// TIA Portal project "Projekt_Serhii_Bodnia" (V19) (continued)

   FOR #forVal := 0 TO 120 DO
       FOR #forVal_2:=0 TO 10 DO
           #rdTimeReturn:=RD_SYS_T(#outputTime);
           #rdTimeReturn := WR_SYS_T(#outputTime);
           #rdTimeReturn := RD_SYS_T(#outputTime);
           #rdTimeReturn := WR_SYS_T(#outputTime);
       END_FOR;
       #SyncVal:= PEEK(area := 16#81,
                      dbNumber := 0,
                      byteOffset := 511);
       IF #SyncVal = #CompVal THEN
          GOTO M_1;
       END_IF;
   END_FOR;
   RETURN;

   M_1:
   POKE(area := 16#81,
        dbNumber := 0,
        byteOffset := 511,
        value := B#16#0);
END_FUNCTION

ORGANIZATION_BLOCK "Main"   // OB1, FBD, ProgramCycle
TITLE = "Main Program Sweep (Cycle)"
{ S7_Optimized_Access := 'TRUE' }
VERSION : 0.1
   VAR_INPUT
      Initial_Call : Bool;   // Initial call of this OB
      Remanence : Bool;   // =True, if remanent data are available
   END_VAR
BEGIN

REGION Network 1: Konnektierungsbaustein für PLC-Lab / Factory IO
   // Im Netzwerk 1 wird der Konnektierungsbaustein für PLC-Lab aufgerufen.
   // Dieser Aufruf darf nicht entfernt werden!
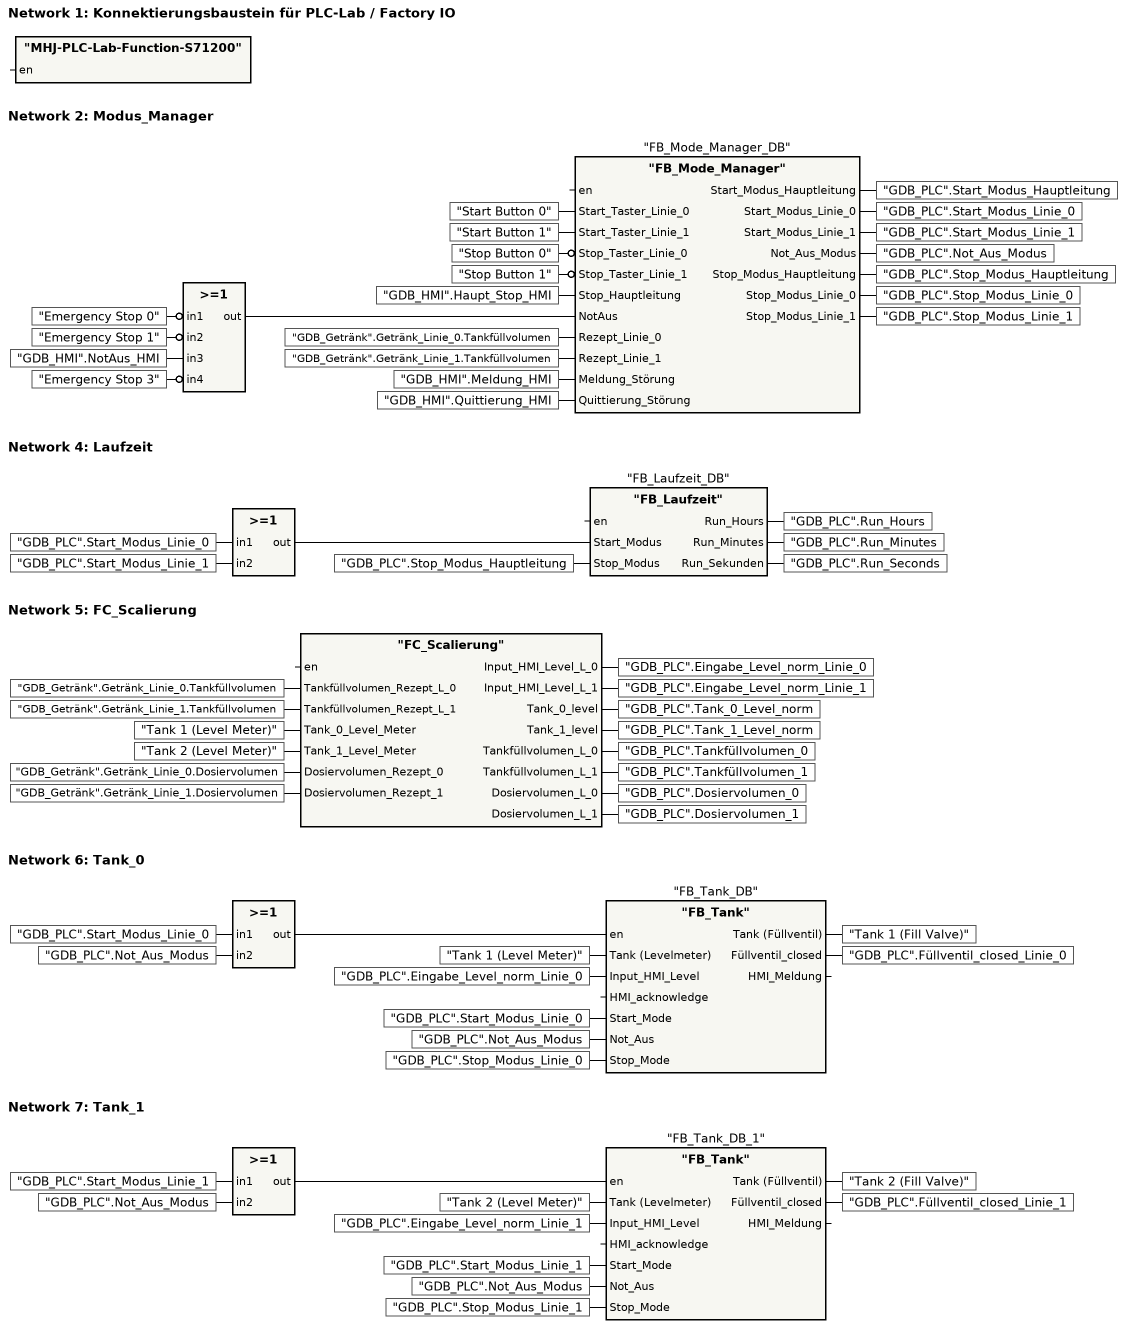
   "MHJ-PLC-Lab-Function-S71200"();
END_REGION

REGION Network 2: Modus_Manager
   "FB_Mode_Manager_DB"(Start_Taster_Linie_0 := "Start Button 0",   // "FB_Mode_Manager"
                        Start_Taster_Linie_1 := "Start Button 1",
                        Stop_Taster_Linie_0 := NOT "Stop Button 0",
                        Stop_Taster_Linie_1 := NOT "Stop Button 1",
                        Stop_Hauptleitung := "GDB_HMI".Haupt_Stop_HMI,
                        NotAus := NOT "Emergency Stop 0" OR NOT "Emergency Stop 1" OR "GDB_HMI".NotAus_HMI OR NOT "Emergency Stop 3",
                        Rezept_Linie_0 := "GDB_Getränk".Getränk_Linie_0.Tankfüllvolumen,
                        Rezept_Linie_1 := "GDB_Getränk".Getränk_Linie_1.Tankfüllvolumen,
                        Meldung_Störung := "GDB_HMI".Meldung_HMI,
                        Quittierung_Störung := "GDB_HMI".Quittierung_HMI,
                        Start_Modus_Hauptleitung => "GDB_PLC".Start_Modus_Hauptleitung,
                        Start_Modus_Linie_0 => "GDB_PLC".Start_Modus_Linie_0,
                        Start_Modus_Linie_1 => "GDB_PLC".Start_Modus_Linie_1,
                        Not_Aus_Modus => "GDB_PLC".Not_Aus_Modus,
                        Stop_Modus_Hauptleitung => "GDB_PLC".Stop_Modus_Hauptleitung,
                        Stop_Modus_Linie_0 => "GDB_PLC".Stop_Modus_Linie_0,
                        Stop_Modus_Linie_1 => "GDB_PLC".Stop_Modus_Linie_1);
END_REGION

REGION Network 3 (SCL): Störung Meldungen
   "GDB_PLC".Störung[0] := "GDB_HMI".Meldung_HMI.%X0;
   "GDB_PLC".Störung[1] := "GDB_HMI".Meldung_HMI.%X1;
   "GDB_PLC".Störung[2] := "GDB_HMI".Meldung_HMI.%X2;
   "GDB_PLC".Störung[3] := "GDB_HMI".Meldung_HMI.%X3;
   "GDB_PLC".Störung[4] := "GDB_HMI".Meldung_HMI.%X4;
   "GDB_PLC".Störung[5] := "GDB_HMI".Meldung_HMI.%X5;
   "GDB_PLC".Störung[6] := "GDB_HMI".Meldung_HMI.%X6;
   "GDB_PLC".Störung[7] := "GDB_HMI".Meldung_HMI.%X7;
   "GDB_PLC".Störung[8] := "GDB_HMI".Meldung_HMI.%X8;
   "GDB_PLC".Störung[9] := "GDB_HMI".Meldung_HMI.%X9;
   "GDB_PLC".Störung[10] := "GDB_HMI".Meldung_HMI.%X10;
   "GDB_PLC".Störung[11] := "GDB_HMI".Meldung_HMI.%X11;
   "GDB_PLC".Störung[12] := "GDB_HMI".Meldung_HMI.%X12;
   "GDB_PLC".Störung[13] := "GDB_HMI".Meldung_HMI.%X13;
   "GDB_PLC".Störung[14] := "GDB_HMI".Meldung_HMI.%X14;
   "GDB_PLC".Störung[15] := "GDB_HMI".Meldung_HMI.%X15;
END_REGION

REGION Network 4: Laufzeit
   "FB_Laufzeit_DB"(Start_Modus := "GDB_PLC".Start_Modus_Linie_0 OR "GDB_PLC".Start_Modus_Linie_1,   // "FB_Laufzeit"
                    Stop_Modus := "GDB_PLC".Stop_Modus_Hauptleitung,
                    Run_Hours => "GDB_PLC".Run_Hours,
                    Run_Minutes => "GDB_PLC".Run_Minutes,
                    Run_Sekunden => "GDB_PLC".Run_Seconds);
END_REGION

REGION Network 5: FC_Scalierung
   "FC_Scalierung"(Tankfüllvolumen_Rezept_L_0 := "GDB_Getränk".Getränk_Linie_0.Tankfüllvolumen,
                   Tankfüllvolumen_Rezept_L_1 := "GDB_Getränk".Getränk_Linie_1.Tankfüllvolumen,
                   Tank_0_Level_Meter := "Tank 1 (Level Meter)",
                   Tank_1_Level_Meter := "Tank 2 (Level Meter)",
                   Dosiervolumen_Rezept_0 := "GDB_Getränk".Getränk_Linie_0.Dosiervolumen,
                   Dosiervolumen_Rezept_1 := "GDB_Getränk".Getränk_Linie_1.Dosiervolumen,
                   Input_HMI_Level_L_0 => "GDB_PLC".Eingabe_Level_norm_Linie_0,
                   Input_HMI_Level_L_1 => "GDB_PLC".Eingabe_Level_norm_Linie_1,
                   Tank_0_level => "GDB_PLC".Tank_0_Level_norm,
                   Tank_1_level => "GDB_PLC".Tank_1_Level_norm,
                   Tankfüllvolumen_L_0 => "GDB_PLC".Tankfüllvolumen_0,
                   Tankfüllvolumen_L_1 => "GDB_PLC".Tankfüllvolumen_1,
                   Dosiervolumen_L_0 => "GDB_PLC".Dosiervolumen_0,
                   Dosiervolumen_L_1 => "GDB_PLC".Dosiervolumen_1);
END_REGION

REGION Network 6: Tank_0
   IF "GDB_PLC".Start_Modus_Linie_0 OR "GDB_PLC".Not_Aus_Modus THEN
       "FB_Tank_DB"("Tank (Levelmeter)" := "Tank 1 (Level Meter)",   // "FB_Tank"
                    Input_HMI_Level := "GDB_PLC".Eingabe_Level_norm_Linie_0,
                    Start_Mode := "GDB_PLC".Start_Modus_Linie_0,
                    Not_Aus := "GDB_PLC".Not_Aus_Modus,
                    Stop_Mode := "GDB_PLC".Stop_Modus_Linie_0,
                    "Tank (Füllventil)" => "Tank 1 (Fill Valve)",
                    Füllventil_closed => "GDB_PLC".Füllventil_closed_Linie_0);
   END_IF;
END_REGION

REGION Network 7: Tank_1
   IF "GDB_PLC".Start_Modus_Linie_1 OR "GDB_PLC".Not_Aus_Modus THEN
       "FB_Tank_DB_1"("Tank (Levelmeter)" := "Tank 2 (Level Meter)",   // "FB_Tank"
                      Input_HMI_Level := "GDB_PLC".Eingabe_Level_norm_Linie_1,
                      Start_Mode := "GDB_PLC".Start_Modus_Linie_1,
                      Not_Aus := "GDB_PLC".Not_Aus_Modus,
                      Stop_Mode := "GDB_PLC".Stop_Modus_Linie_1,
                      "Tank (Füllventil)" => "Tank 2 (Fill Valve)",
                      Füllventil_closed => "GDB_PLC".Füllventil_closed_Linie_1);
   END_IF;
END_REGION

REGION Network 8: Abfüllmaschine_Band_0
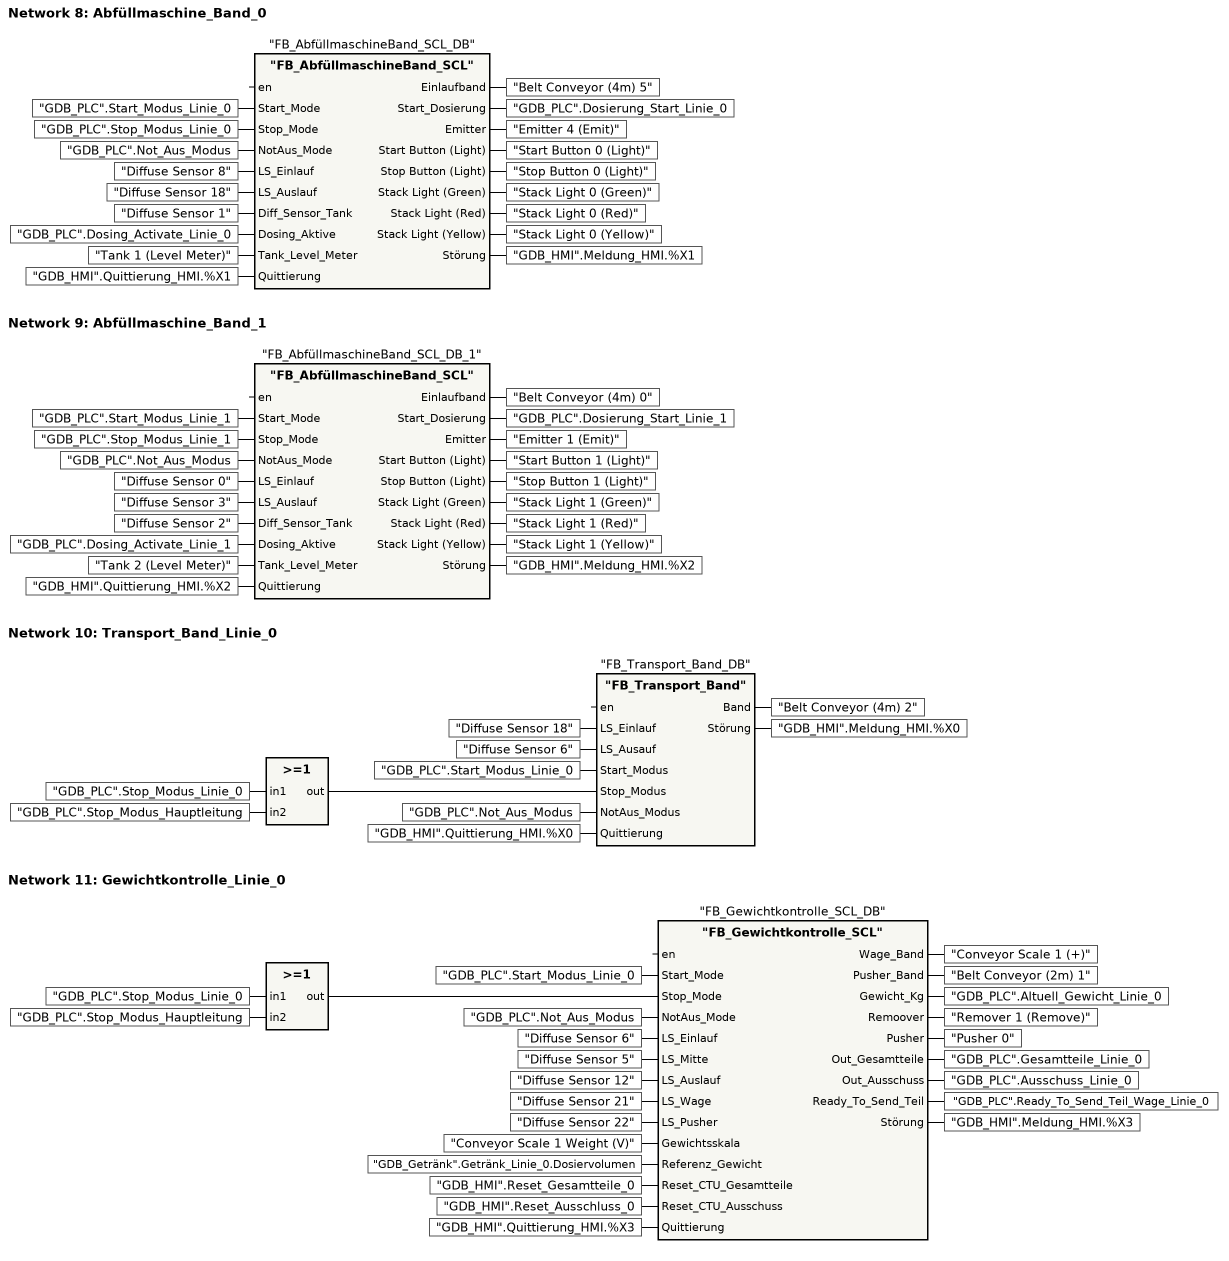
   "FB_AbfüllmaschineBand_SCL_DB"(Start_Mode := "GDB_PLC".Start_Modus_Linie_0,   // "FB_AbfüllmaschineBand_SCL"
                           Stop_Mode := "GDB_PLC".Stop_Modus_Linie_0,
                           NotAus_Mode := "GDB_PLC".Not_Aus_Modus,
                           LS_Einlauf := "Diffuse Sensor 8",
                           LS_Auslauf := "Diffuse Sensor 18",
                           Diff_Sensor_Tank := "Diffuse Sensor 1",
                           Dosing_Aktive := "GDB_PLC".Dosing_Activate_Linie_0,
                           Tank_Level_Meter := "Tank 1 (Level Meter)",
                           Quittierung := "GDB_HMI".Quittierung_HMI.%X1,
                           Einlaufband => "Belt Conveyor (4m) 5",
                           Start_Dosierung => "GDB_PLC".Dosierung_Start_Linie_0,
                           Emitter => "Emitter 4 (Emit)",
                           "Start Button (Light)" => "Start Button 0 (Light)",
                           "Stop Button (Light)" => "Stop Button 0 (Light)",
                           "Stack Light (Green)" => "Stack Light 0 (Green)",
                           "Stack Light (Red)" => "Stack Light 0 (Red)",
                           "Stack Light (Yellow)" => "Stack Light 0 (Yellow)",
                           Störung => "GDB_HMI".Meldung_HMI.%X1);
END_REGION

REGION Network 9: Abfüllmaschine_Band_1
   "FB_AbfüllmaschineBand_SCL_DB_1"(Start_Mode := "GDB_PLC".Start_Modus_Linie_1,   // "FB_AbfüllmaschineBand_SCL"
                           Stop_Mode := "GDB_PLC".Stop_Modus_Linie_1,
                           NotAus_Mode := "GDB_PLC".Not_Aus_Modus,
                           LS_Einlauf := "Diffuse Sensor 0",
                           LS_Auslauf := "Diffuse Sensor 3",
                           Diff_Sensor_Tank := "Diffuse Sensor 2",
                           Dosing_Aktive := "GDB_PLC".Dosing_Activate_Linie_1,
                           Tank_Level_Meter := "Tank 2 (Level Meter)",
                           Quittierung := "GDB_HMI".Quittierung_HMI.%X2,
                           Einlaufband => "Belt Conveyor (4m) 0",
                           Start_Dosierung => "GDB_PLC".Dosierung_Start_Linie_1,
                           Emitter => "Emitter 1 (Emit)",
                           "Start Button (Light)" => "Start Button 1 (Light)",
                           "Stop Button (Light)" => "Stop Button 1 (Light)",
                           "Stack Light (Green)" => "Stack Light 1 (Green)",
                           "Stack Light (Red)" => "Stack Light 1 (Red)",
                           "Stack Light (Yellow)" => "Stack Light 1 (Yellow)",
                           Störung => "GDB_HMI".Meldung_HMI.%X2);
END_REGION

REGION Network 10: Transport_Band_Linie_0
   "FB_Transport_Band_DB"(LS_Einlauf := "Diffuse Sensor 18",   // "FB_Transport_Band"
                          LS_Ausauf := "Diffuse Sensor 6",
                          Start_Modus := "GDB_PLC".Start_Modus_Linie_0,
                          Stop_Modus := "GDB_PLC".Stop_Modus_Linie_0 OR "GDB_PLC".Stop_Modus_Hauptleitung,
                          NotAus_Modus := "GDB_PLC".Not_Aus_Modus,
                          Quittierung := "GDB_HMI".Quittierung_HMI.%X0,
                          Band => "Belt Conveyor (4m) 2",
                          Störung => "GDB_HMI".Meldung_HMI.%X0);
END_REGION

REGION Network 11: Gewichtkontrolle_Linie_0
   "FB_Gewichtkontrolle_SCL_DB"(Start_Mode := "GDB_PLC".Start_Modus_Linie_0,   // "FB_Gewichtkontrolle_SCL"
                           Stop_Mode := "GDB_PLC".Stop_Modus_Linie_0 OR "GDB_PLC".Stop_Modus_Hauptleitung,
                           NotAus_Mode := "GDB_PLC".Not_Aus_Modus,
                           LS_Einlauf := "Diffuse Sensor 6",
                           LS_Mitte := "Diffuse Sensor 5",
                           LS_Auslauf := "Diffuse Sensor 12",
                           LS_Wage := "Diffuse Sensor 21",
                           LS_Pusher := "Diffuse Sensor 22",
                           Gewichtsskala := "Conveyor Scale 1 Weight (V)",
                           Referenz_Gewicht := "GDB_Getränk".Getränk_Linie_0.Dosiervolumen,
                           Reset_CTU_Gesamtteile := "GDB_HMI".Reset_Gesamtteile_0,
                           Reset_CTU_Ausschuss := "GDB_HMI".Reset_Ausschluss_0,
                           Quittierung := "GDB_HMI".Quittierung_HMI.%X3,
                           Wage_Band => "Conveyor Scale 1 (+)",
                           Pusher_Band => "Belt Conveyor (2m) 1",
                           Gewicht_Kg => "GDB_PLC".Altuell_Gewicht_Linie_0,
                           Remoover => "Remover 1 (Remove)",
                           Pusher => "Pusher 0",
                           Out_Gesamtteile => "GDB_PLC".Gesamtteile_Linie_0,
                           Out_Ausschuss => "GDB_PLC".Ausschuss_Linie_0,
                           Ready_To_Send_Teil => "GDB_PLC".Ready_To_Send_Teil_Wage_Linie_0,
                           Störung => "GDB_HMI".Meldung_HMI.%X3);
END_REGION

REGION Network 12: Gewichtkontrolle_Linie_1
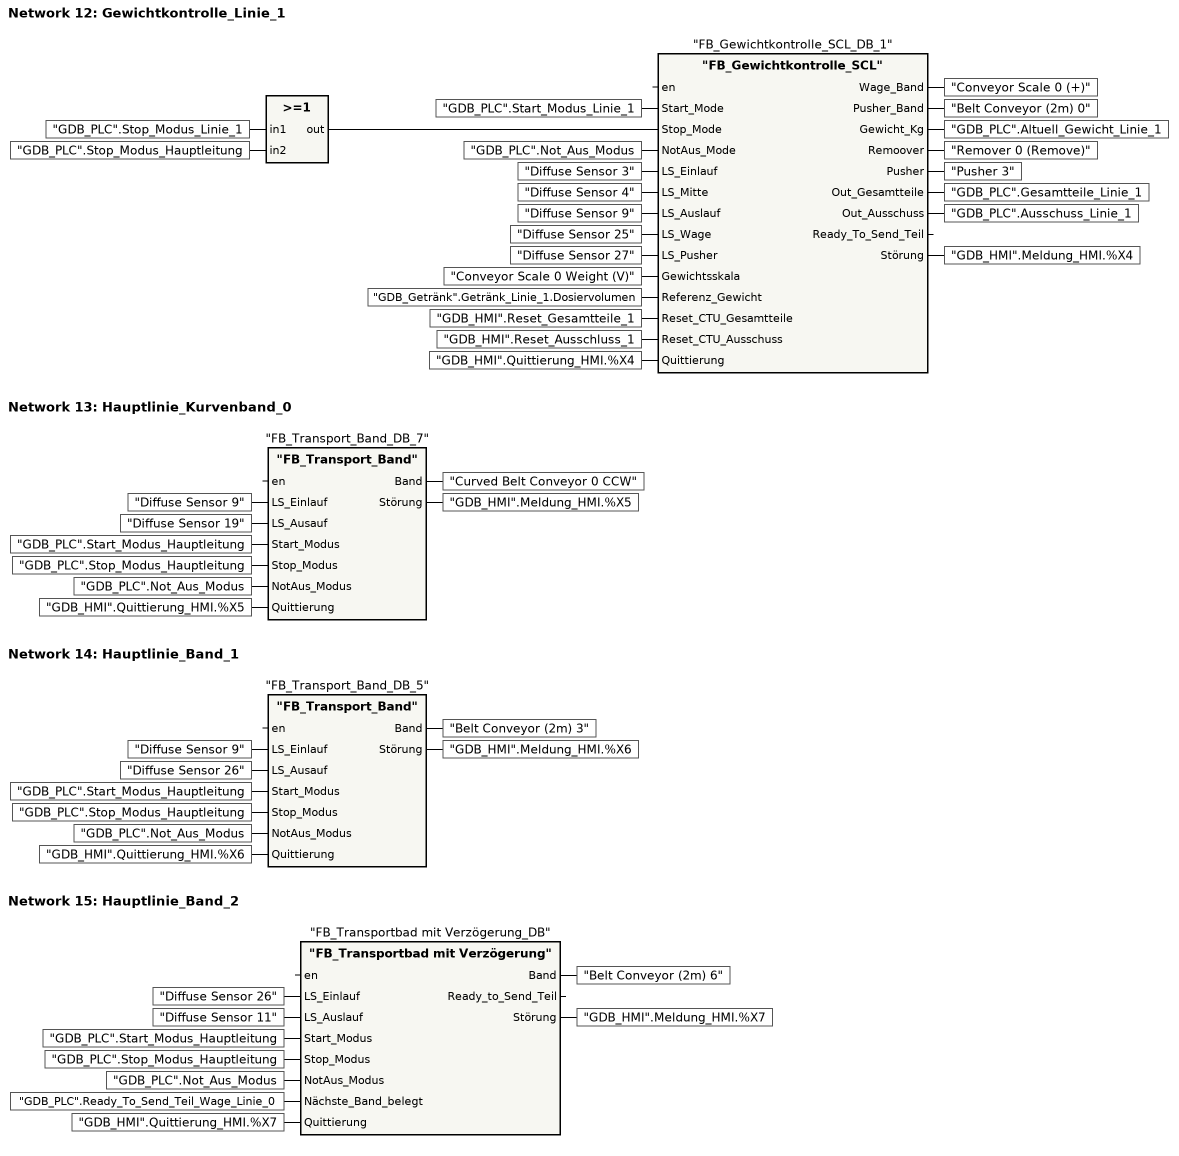
   "FB_Gewichtkontrolle_SCL_DB_1"(Start_Mode := "GDB_PLC".Start_Modus_Linie_1,   // "FB_Gewichtkontrolle_SCL"
                           Stop_Mode := "GDB_PLC".Stop_Modus_Linie_1 OR "GDB_PLC".Stop_Modus_Hauptleitung,
                           NotAus_Mode := "GDB_PLC".Not_Aus_Modus,
                           LS_Einlauf := "Diffuse Sensor 3",
                           LS_Mitte := "Diffuse Sensor 4",
                           LS_Auslauf := "Diffuse Sensor 9",
                           LS_Wage := "Diffuse Sensor 25",
                           LS_Pusher := "Diffuse Sensor 27",
                           Gewichtsskala := "Conveyor Scale 0 Weight (V)",
                           Referenz_Gewicht := "GDB_Getränk".Getränk_Linie_1.Dosiervolumen,
                           Reset_CTU_Gesamtteile := "GDB_HMI".Reset_Gesamtteile_1,
                           Reset_CTU_Ausschuss := "GDB_HMI".Reset_Ausschluss_1,
                           Quittierung := "GDB_HMI".Quittierung_HMI.%X4,
                           Wage_Band => "Conveyor Scale 0 (+)",
                           Pusher_Band => "Belt Conveyor (2m) 0",
                           Gewicht_Kg => "GDB_PLC".Altuell_Gewicht_Linie_1,
                           Remoover => "Remover 0 (Remove)",
                           Pusher => "Pusher 3",
                           Out_Gesamtteile => "GDB_PLC".Gesamtteile_Linie_1,
                           Out_Ausschuss => "GDB_PLC".Ausschuss_Linie_1,
                           Störung => "GDB_HMI".Meldung_HMI.%X4);
END_REGION

REGION Network 13: Hauptlinie_Kurvenband_0
   "FB_Transport_Band_DB_7"(LS_Einlauf := "Diffuse Sensor 9",   // "FB_Transport_Band"
                           LS_Ausauf := "Diffuse Sensor 19",
                           Start_Modus := "GDB_PLC".Start_Modus_Hauptleitung,
                           Stop_Modus := "GDB_PLC".Stop_Modus_Hauptleitung,
                           NotAus_Modus := "GDB_PLC".Not_Aus_Modus,
                           Quittierung := "GDB_HMI".Quittierung_HMI.%X5,
                           Band => "Curved Belt Conveyor 0 CCW",
                           Störung => "GDB_HMI".Meldung_HMI.%X5);
END_REGION

REGION Network 14: Hauptlinie_Band_1
   "FB_Transport_Band_DB_5"(LS_Einlauf := "Diffuse Sensor 9",   // "FB_Transport_Band"
                           LS_Ausauf := "Diffuse Sensor 26",
                           Start_Modus := "GDB_PLC".Start_Modus_Hauptleitung,
                           Stop_Modus := "GDB_PLC".Stop_Modus_Hauptleitung,
                           NotAus_Modus := "GDB_PLC".Not_Aus_Modus,
                           Quittierung := "GDB_HMI".Quittierung_HMI.%X6,
                           Band => "Belt Conveyor (2m) 3",
                           Störung => "GDB_HMI".Meldung_HMI.%X6);
END_REGION

REGION Network 15: Hauptlinie_Band_2
   "FB_Transportbad mit Verzögerung_DB"(LS_Einlauf := "Diffuse Sensor 26",   // "FB_Transportbad mit Verzögerung"
                           LS_Auslauf := "Diffuse Sensor 11",
                           Start_Modus := "GDB_PLC".Start_Modus_Hauptleitung,
                           Stop_Modus := "GDB_PLC".Stop_Modus_Hauptleitung,
                           NotAus_Modus := "GDB_PLC".Not_Aus_Modus,
                           Nächste_Band_belegt := "GDB_PLC".Ready_To_Send_Teil_Wage_Linie_0,
                           Quittierung := "GDB_HMI".Quittierung_HMI.%X7,
                           Band => "Belt Conveyor (2m) 6",
                           Störung => "GDB_HMI".Meldung_HMI.%X7);
END_REGION

REGION Network 16: Hauptlinie_T - Band_3
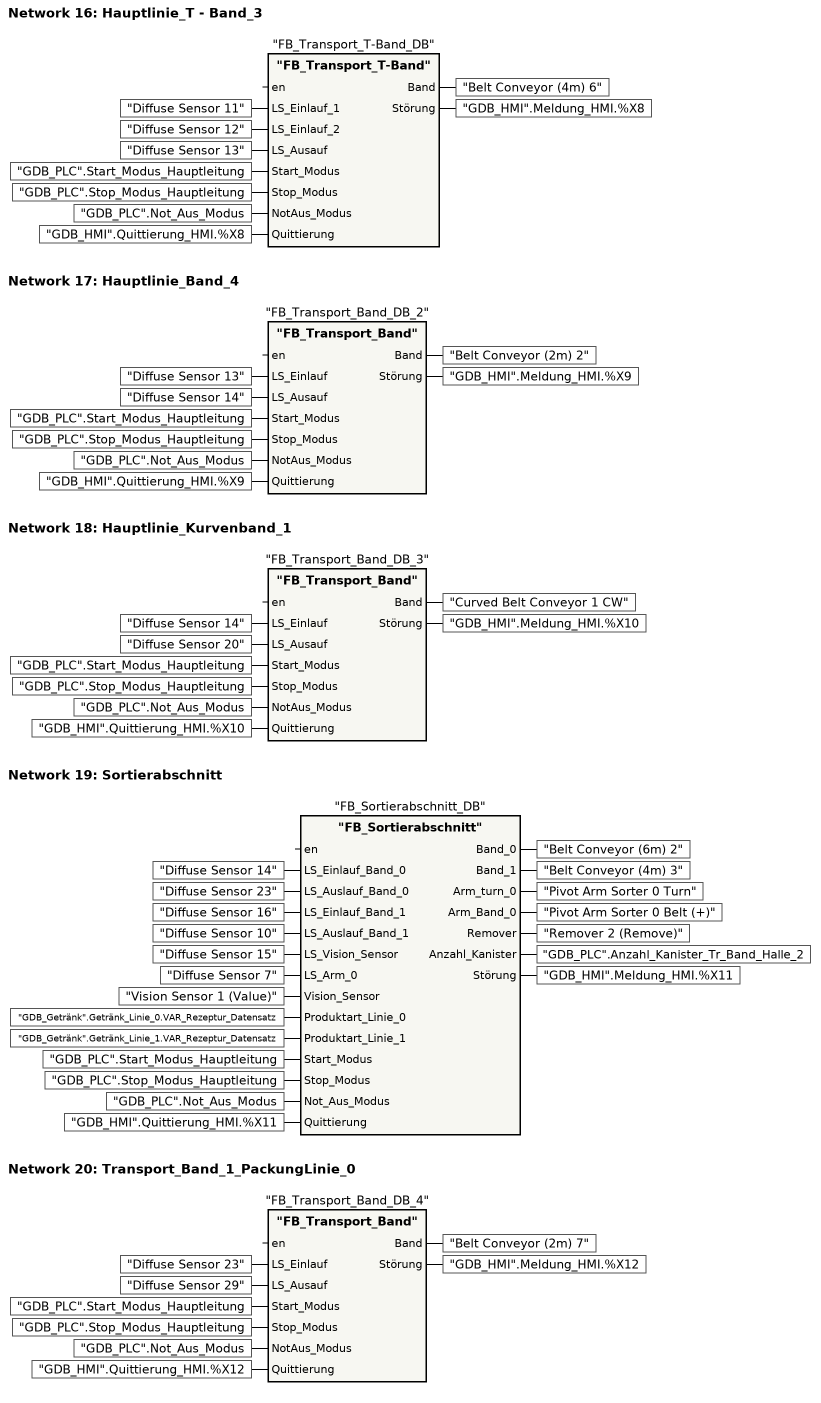
   "FB_Transport_T-Band_DB"(LS_Einlauf_1 := "Diffuse Sensor 11",   // "FB_Transport_T-Band"
                           LS_Einlauf_2 := "Diffuse Sensor 12",
                           LS_Ausauf := "Diffuse Sensor 13",
                           Start_Modus := "GDB_PLC".Start_Modus_Hauptleitung,
                           Stop_Modus := "GDB_PLC".Stop_Modus_Hauptleitung,
                           NotAus_Modus := "GDB_PLC".Not_Aus_Modus,
                           Quittierung := "GDB_HMI".Quittierung_HMI.%X8,
                           Band => "Belt Conveyor (4m) 6",
                           Störung => "GDB_HMI".Meldung_HMI.%X8);
END_REGION

REGION Network 17: Hauptlinie_Band_4
   "FB_Transport_Band_DB_2"(LS_Einlauf := "Diffuse Sensor 13",   // "FB_Transport_Band"
                           LS_Ausauf := "Diffuse Sensor 14",
                           Start_Modus := "GDB_PLC".Start_Modus_Hauptleitung,
                           Stop_Modus := "GDB_PLC".Stop_Modus_Hauptleitung,
                           NotAus_Modus := "GDB_PLC".Not_Aus_Modus,
                           Quittierung := "GDB_HMI".Quittierung_HMI.%X9,
                           Band => "Belt Conveyor (2m) 2",
                           Störung => "GDB_HMI".Meldung_HMI.%X9);
END_REGION

REGION Network 18: Hauptlinie_Kurvenband_1
   "FB_Transport_Band_DB_3"(LS_Einlauf := "Diffuse Sensor 14",   // "FB_Transport_Band"
                           LS_Ausauf := "Diffuse Sensor 20",
                           Start_Modus := "GDB_PLC".Start_Modus_Hauptleitung,
                           Stop_Modus := "GDB_PLC".Stop_Modus_Hauptleitung,
                           NotAus_Modus := "GDB_PLC".Not_Aus_Modus,
                           Quittierung := "GDB_HMI".Quittierung_HMI.%X10,
                           Band => "Curved Belt Conveyor 1 CW",
                           Störung => "GDB_HMI".Meldung_HMI.%X10);
END_REGION

REGION Network 19: Sortierabschnitt
   "FB_Sortierabschnitt_DB"(LS_Einlauf_Band_0 := "Diffuse Sensor 14",   // "FB_Sortierabschnitt"
                           LS_Auslauf_Band_0 := "Diffuse Sensor 23",
                           LS_Einlauf_Band_1 := "Diffuse Sensor 16",
                           LS_Auslauf_Band_1 := "Diffuse Sensor 10",
                           LS_Vision_Sensor := "Diffuse Sensor 15",
                           LS_Arm_0 := "Diffuse Sensor 7",
                           Vision_Sensor := "Vision Sensor 1 (Value)",
                           Produktart_Linie_0 := "GDB_Getränk".Getränk_Linie_0.VAR_Rezeptur_Datensatz,
                           Produktart_Linie_1 := "GDB_Getränk".Getränk_Linie_1.VAR_Rezeptur_Datensatz,
                           Start_Modus := "GDB_PLC".Start_Modus_Hauptleitung,
                           Stop_Modus := "GDB_PLC".Stop_Modus_Hauptleitung,
                           Not_Aus_Modus := "GDB_PLC".Not_Aus_Modus,
                           Quittierung := "GDB_HMI".Quittierung_HMI.%X11,
                           Band_0 => "Belt Conveyor (6m) 2",
                           Band_1 => "Belt Conveyor (4m) 3",
                           Arm_turn_0 => "Pivot Arm Sorter 0 Turn",
                           Arm_Band_0 => "Pivot Arm Sorter 0 Belt (+)",
                           Remover => "Remover 2 (Remove)",
                           Anzahl_Kanister => "GDB_PLC".Anzahl_Kanister_Tr_Band_Halle_2,
                           Störung => "GDB_HMI".Meldung_HMI.%X11);
END_REGION

REGION Network 20: Transport_Band_1_PackungLinie_0
   "FB_Transport_Band_DB_4"(LS_Einlauf := "Diffuse Sensor 23",   // "FB_Transport_Band"
                           LS_Ausauf := "Diffuse Sensor 29",
                           Start_Modus := "GDB_PLC".Start_Modus_Hauptleitung,
                           Stop_Modus := "GDB_PLC".Stop_Modus_Hauptleitung,
                           NotAus_Modus := "GDB_PLC".Not_Aus_Modus,
                           Quittierung := "GDB_HMI".Quittierung_HMI.%X12,
                           Band => "Belt Conveyor (2m) 7",
                           Störung => "GDB_HMI".Meldung_HMI.%X12);
END_REGION

REGION Network 21: Transport_Band_2_PackungLinie_0
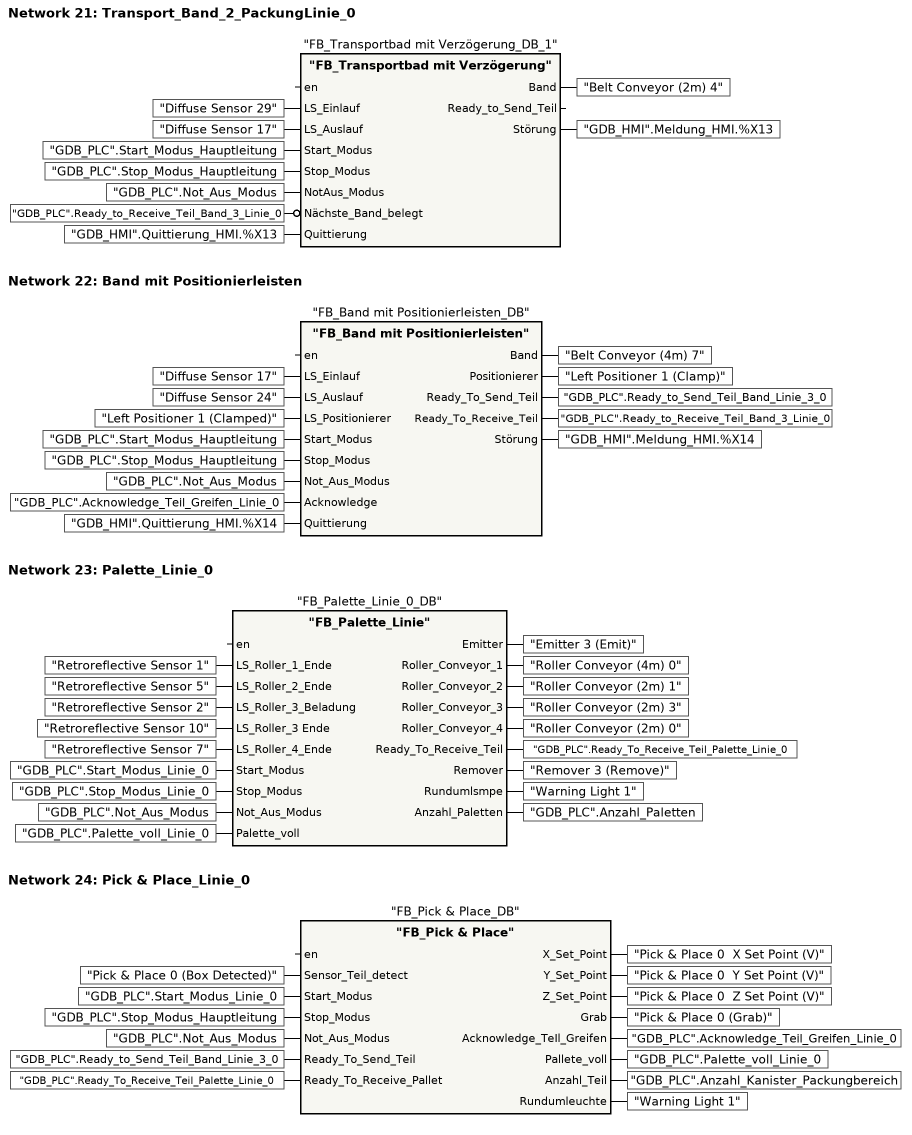
   "FB_Transportbad mit Verzögerung_DB_1"(LS_Einlauf := "Diffuse Sensor 29",   // "FB_Transportbad mit Verzögerung"
                           LS_Auslauf := "Diffuse Sensor 17",
                           Start_Modus := "GDB_PLC".Start_Modus_Hauptleitung,
                           Stop_Modus := "GDB_PLC".Stop_Modus_Hauptleitung,
                           NotAus_Modus := "GDB_PLC".Not_Aus_Modus,
                           Nächste_Band_belegt := NOT "GDB_PLC".Ready_to_Receive_Teil_Band_3_Linie_0,
                           Quittierung := "GDB_HMI".Quittierung_HMI.%X13,
                           Band => "Belt Conveyor (2m) 4",
                           Störung => "GDB_HMI".Meldung_HMI.%X13);
END_REGION

REGION Network 22: Band mit Positionierleisten
   "FB_Band mit Positionierleisten_DB"(LS_Einlauf := "Diffuse Sensor 17",   // "FB_Band mit Positionierleisten"
                           LS_Auslauf := "Diffuse Sensor 24",
                           LS_Positionierer := "Left Positioner 1 (Clamped)",
                           Start_Modus := "GDB_PLC".Start_Modus_Hauptleitung,
                           Stop_Modus := "GDB_PLC".Stop_Modus_Hauptleitung,
                           Not_Aus_Modus := "GDB_PLC".Not_Aus_Modus,
                           Acknowledge := "GDB_PLC".Acknowledge_Teil_Greifen_Linie_0,
                           Quittierung := "GDB_HMI".Quittierung_HMI.%X14,
                           Band => "Belt Conveyor (4m) 7",
                           Positionierer => "Left Positioner 1 (Clamp)",
                           Ready_To_Send_Teil => "GDB_PLC".Ready_to_Send_Teil_Band_Linie_3_0,
                           Ready_To_Receive_Teil => "GDB_PLC".Ready_to_Receive_Teil_Band_3_Linie_0,
                           Störung => "GDB_HMI".Meldung_HMI.%X14);
END_REGION

REGION Network 23: Palette_Linie_0
   "FB_Palette_Linie_0_DB"(LS_Roller_1_Ende := "Retroreflective Sensor 1",   // "FB_Palette_Linie"
                           LS_Roller_2_Ende := "Retroreflective Sensor 5",
                           LS_Roller_3_Beladung := "Retroreflective Sensor 2",
                           "LS_Roller_3 Ende" := "Retroreflective Sensor 10",
                           LS_Roller_4_Ende := "Retroreflective Sensor 7",
                           Start_Modus := "GDB_PLC".Start_Modus_Linie_0,
                           Stop_Modus := "GDB_PLC".Stop_Modus_Linie_0,
                           Not_Aus_Modus := "GDB_PLC".Not_Aus_Modus,
                           Palette_voll := "GDB_PLC".Palette_voll_Linie_0,
                           Emitter => "Emitter 3 (Emit)",
                           Roller_Conveyor_1 => "Roller Conveyor (4m) 0",
                           Roller_Conveyor_2 => "Roller Conveyor (2m) 1",
                           Roller_Conveyor_3 => "Roller Conveyor (2m) 3",
                           Roller_Conveyor_4 => "Roller Conveyor (2m) 0",
                           Ready_To_Receive_Teil => "GDB_PLC".Ready_To_Receive_Teil_Palette_Linie_0,
                           Remover => "Remover 3 (Remove)",
                           Rundumlsmpe => "Warning Light 1",
                           Anzahl_Paletten => "GDB_PLC".Anzahl_Paletten);
END_REGION

REGION Network 24: Pick & Place_Linie_0
   "FB_Pick & Place_DB"(Sensor_Teil_detect := "Pick & Place 0 (Box Detected)",   // "FB_Pick & Place"
                        Start_Modus := "GDB_PLC".Start_Modus_Linie_0,
                        Stop_Modus := "GDB_PLC".Stop_Modus_Hauptleitung,
                        Not_Aus_Modus := "GDB_PLC".Not_Aus_Modus,
                        Ready_To_Send_Teil := "GDB_PLC".Ready_to_Send_Teil_Band_Linie_3_0,
                        Ready_To_Receive_Pallet := "GDB_PLC".Ready_To_Receive_Teil_Palette_Linie_0,
                        X_Set_Point => "Pick & Place 0  X Set Point (V)",
                        Y_Set_Point => "Pick & Place 0  Y Set Point (V)",
                        Z_Set_Point => "Pick & Place 0  Z Set Point (V)",
                        Grab => "Pick & Place 0 (Grab)",
                        Acknowledge_TeIl_Greifen => "GDB_PLC".Acknowledge_Teil_Greifen_Linie_0,
                        Pallete_voll => "GDB_PLC".Palette_voll_Linie_0,
                        Anzahl_Teil => "GDB_PLC".Anzahl_Kanister_Packungbereich,
                        Rundumleuchte => "Warning Light 1");
END_REGION
END_ORGANIZATION_BLOCK

ORGANIZATION_BLOCK "Cyclic interrupt"   // OB30, FBD, CyclicInterrupt
{ S7_Optimized_Access := 'TRUE' }
VERSION : 0.1
   VAR_INPUT
      Initial_Call : Bool;   // Initial call of this OB
      Event_Count : Int;   // Events discarded
   END_VAR
BEGIN

REGION Network 1: Dose_Control_Linie_0
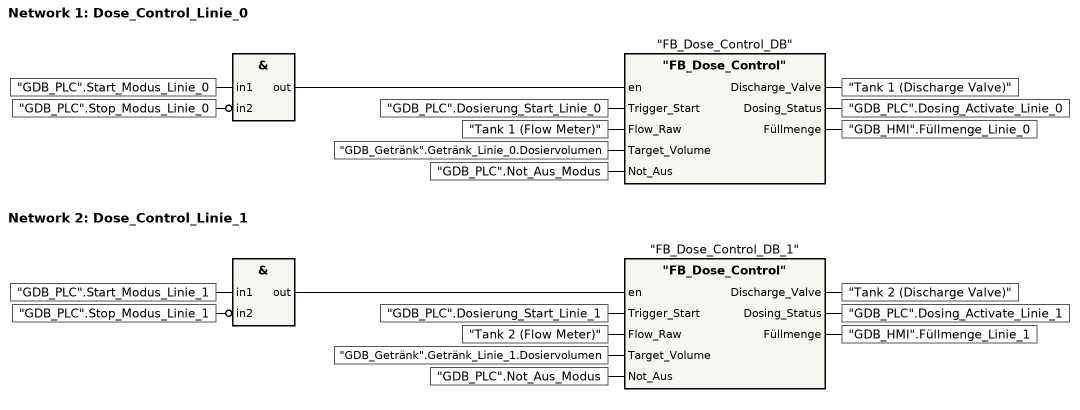
   IF "GDB_PLC".Start_Modus_Linie_0 AND NOT "GDB_PLC".Stop_Modus_Linie_0 THEN
       "FB_Dose_Control_DB"(Trigger_Start := "GDB_PLC".Dosierung_Start_Linie_0,   // "FB_Dose_Control"
                            Flow_Raw := "Tank 1 (Flow Meter)",
                            Target_Volume := "GDB_Getränk".Getränk_Linie_0.Dosiervolumen,
                            Not_Aus := "GDB_PLC".Not_Aus_Modus,
                            Discharge_Valve => "Tank 1 (Discharge Valve)",
                            Dosing_Status => "GDB_PLC".Dosing_Activate_Linie_0,
                            Füllmenge => "GDB_HMI".Füllmenge_Linie_0);
   END_IF;
END_REGION

